
       FOR #Idx2 := 1 TO #Idx1 + 1 DO
           IF #ArrayTemp[#Idx2].Position > #MaxVal THEN
               #MaxVal := #ArrayTemp[#Idx2].Position;
               #MaxCarr := #ArrayTemp[#Idx2].CarrierNumber;
               #MaxIdx1 := #Idx2;
           END_IF;
       END_FOR;
       IF #MaxIdx1 > #Idx1 THEN
           #ArrayTemp[#MaxIdx1].Position := #ArrayTemp[#Idx1].Position;
           #ArrayTemp[#MaxIdx1].CarrierNumber := #ArrayTemp[#Idx1].CarrierNumber;
           #ArrayTemp[#Idx1].Position := #MaxVal;
           #ArrayTemp[#Idx1].CarrierNumber := #MaxCarr;

       END_IF;

   END_FOR;
   #ZonePositionArrayOut := #ArrayTemp;
END_FUNCTION

FUNCTION "FC107_FindLastZnPos" : Void   // FC107, SCL
{ S7_Optimized_Access := 'FALSE' }
VERSION : 0.1
   VAR_INPUT
      Zone : Int;
      TotalPosition : Int;
   END_VAR
   VAR_OUTPUT
      LastCarrierZnPos : Word;
   END_VAR
   VAR_TEMP
      ZnPosCounter : Int;
      ZoneFound : Word;
      CarrierCounter : Int;
      SortArrayIndex : Int;
      ArrayIndex : Int;
      Idx1 : Int;
      MaxVal : Int;
      MaxIdx1 : Int;
      Max : Int;
      Idx2 : Int;
      SelectionSort : Int;
   END_VAR
BEGIN
       #ZnPosCounter := #TotalPosition;
       WHILE #ZnPosCounter >= 1 DO

           IF "EMS".Zone[#Zone].CarrierZnStatus[#ZnPosCounter].CarrierNumber <> 0 THEN
               ;
               #LastCarrierZnPos := #ZnPosCounter;
               RETURN;
           END_IF;
           #ZnPosCounter := #ZnPosCounter - 1;
       END_WHILE;
END_FUNCTION

FUNCTION "FC108_FindCarrierZNPos" : Void   // FC108, SCL
{ S7_Optimized_Access := 'FALSE' }
VERSION : 0.1
   VAR_INPUT
      Carrier : Word;
      Zone : Int;
      TotalPosition : Int;
   END_VAR
   VAR_OUTPUT
      CarrierZnPos : Word;
   END_VAR
   VAR_TEMP
      ZnPosCounter : Int;
      ZoneFound : Word;
      CarrierCounter : Int;
      SortArrayIndex : Int;
      ArrayIndex : Int;
      Idx1 : Int;
      MaxVal : Int;
      MaxIdx1 : Int;
      Max : Int;
      Idx2 : Int;
      SelectionSort : Int;
   END_VAR
BEGIN
   //[***********************************************************************************NO EDITS*******************************************************************************************************]
   //FC204 - Find Carrier Zone Position
   //Single loop Counter finds which #Zone Position. Zone Position is determined BY Value OF Max Carriers defined in  #Carrier is located based on #Zone Start Position AND End Position AND
   //records the result in the system "EMS" DB FOR each Zone and the results stored in the EMS.Zone[Zone].CarrierZnStatus[1 thru Max Carriers in Zone].Carrier Number
   //***************************************************************************************************************************************************************************************************   

       #ZnPosCounter := 1;
       FOR #ZnPosCounter := 1 TO #TotalPosition DO
           ;
           IF "EMS".Zone[#Zone].CarrierZnStatus[#ZnPosCounter].CarrierNumber = #Carrier THEN;
               ;
               #CarrierZnPos := #ZnPosCounter;
           END_IF;
       END_FOR;
END_FUNCTION

FUNCTION "FC109_FindDuplicateCarrier" : Void   // FC109, SCL
{ S7_Optimized_Access := 'TRUE' }
VERSION : 0.1
   VAR_INPUT
      Carrier : Array[0..99] of "UDT_CarrierStructure";
      TotalCarriers : Int;
   END_VAR
   VAR_OUTPUT
      DuplicateFound : Bool;
      DuplicateCarrierNumber : Word;
      FirstDuplicatePosition : Word;
      SecondDuplicate : Word;
   END_VAR
   VAR_TEMP
      CarrierFindCnt : Int;
      temp1 : Int;
      CarrierCounter : Int;
      CarrierFindArray : Array[0..99] of "UDT_CarrierStructure";
   END_VAR
BEGIN
   //Sorts Carriers in Called Zone TO place in correct sequence within  Zone. Zones are divided into position based on MaxCarriers allowed in Zone as set in the Zone setup function block.


   #DuplicateFound := FALSE;
   #CarrierCounter := 1;
   #CarrierFindCnt := 1;
   #CarrierFindArray := #Carrier;
   FOR #CarrierFindCnt := 1 TO #TotalCarriers DO
       ;
       WHILE #CarrierCounter <= #TotalCarriers DO
           ;
           IF #Carrier[#CarrierCounter].SDC_IN.CarrierNumber = #CarrierFindArray[#CarrierFindCnt].SDC_IN.CarrierNumber AND #CarrierCounter <> #CarrierFindCnt AND #Carrier[#CarrierCounter].SDC_IN.CarrierNumber <> 0 THEN
               #DuplicateFound := TRUE;
               #FirstDuplicatePosition:= #Carrier[#CarrierCounter].SDC_IN.CarrierPosition;
               #SecondDuplicate := #Carrier[#CarrierFindCnt].SDC_IN.CarrierPosition;
               #DuplicateCarrierNumber := #CarrierFindArray[#CarrierFindCnt].SDC_IN.CarrierNumber;
               RETURN;
           END_IF;
           #CarrierCounter := #CarrierCounter + 1;
       END_WHILE;

       #CarrierCounter := 1;
   END_FOR;
END_FUNCTION

FUNCTION "FC110_HMIZonePosTracking" : Void   // FC110, SCL
{ S7_Optimized_Access := 'FALSE' }
VERSION : 0.1
   VAR_INPUT
      Zone : Int;
      TotalZones : Int;
      TotalCarriers : Int;
      MaxCarrierPosns : Int;
   END_VAR
   VAR_OUTPUT
      HMIZonePositionDisplay : Array[1..20] of "UDT_HMIZonePositionStructure";
   END_VAR
   VAR_TEMP
      PositionCounter : Int;
      ZoneFound : Word;
      CarrierCounter : Int;
      ZouneFound : Int;
   END_VAR
BEGIN

       FOR #PositionCounter := 1 TO #MaxCarrierPosns BY 1 DO
           FOR #CarrierCounter := 1 TO #TotalCarriers BY 1 DO
               ;
               IF "EMS".Carrier[#CarrierCounter].Position >= "EMS".Zone[#Zone].HMIZonePositions[#PositionCounter].ZonePosition AND
                   "EMS".Carrier[#CarrierCounter].Position < "EMS".Zone[#Zone].HMIZonePositions[#PositionCounter + 1].ZonePosition
               THEN
                   #HMIZonePositionDisplay[#PositionCounter].CarrierNumber := #CarrierCounter;
                   #HMIZonePositionDisplay[#PositionCounter].CarrierPosition := "EMS".Carrier[#CarrierCounter].Position;
                   #HMIZonePositionDisplay[#PositionCounter].Faulted := "EMS".Carrier[#CarrierCounter].Faulted;
                   EXIT;
               ELSE
                   ;
                   #HMIZonePositionDisplay[#PositionCounter].CarrierNumber := 0;
                   #HMIZonePositionDisplay[#PositionCounter].CarrierPosition := 0;
                   #HMIZonePositionDisplay[#PositionCounter].Faulted := 0;
               END_IF;
               "FC206CarrierLoop" := #CarrierCounter;
           END_FOR;
       "FC206PositionLoop" := #PositionCounter;
   END_FOR;
END_FUNCTION

FUNCTION "FC111_HMI_Status" : Void   // FC111, LAD
{ S7_Optimized_Access := 'TRUE' }
VERSION : 0.1
BEGIN

REGION Network 1
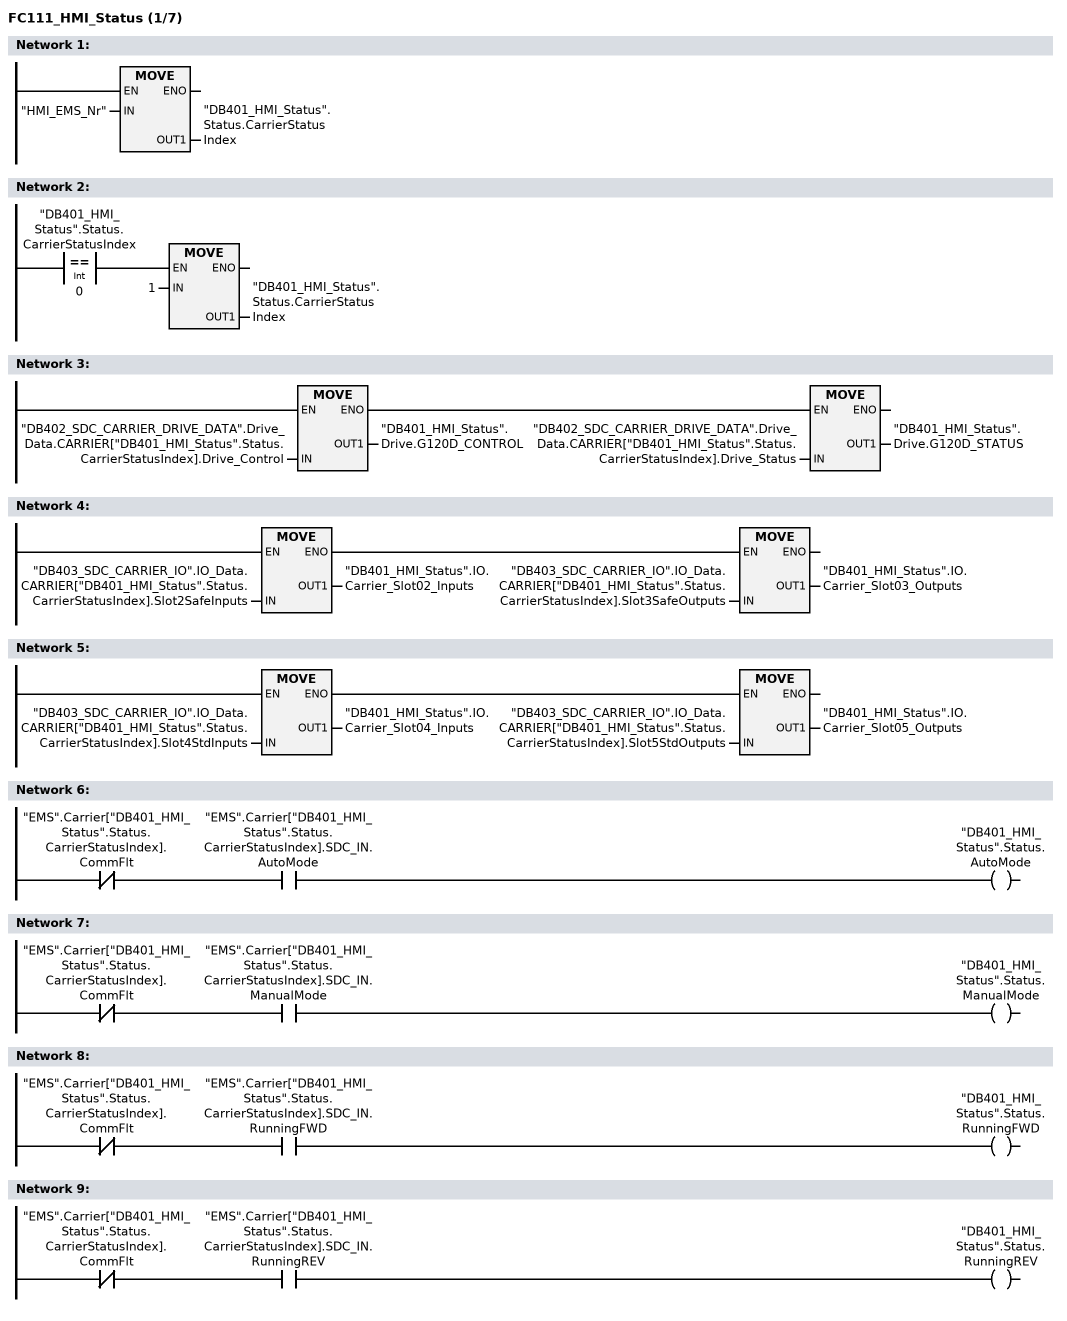
   RUNG wire#powerrail
      Move(in := "HMI_EMS_Nr", out1 => "DB401_HMI_Status".Status.CarrierStatusIndex)
   END_RUNG
   // the same network as SCL:
   "DB401_HMI_Status".Status.CarrierStatusIndex := "HMI_EMS_Nr";
END_REGION

REGION Network 2
   RUNG wire#powerrail
      { S7_Templates := "SrcType := Int" } EQ_Contact(in1 := "DB401_HMI_Status".Status.CarrierStatusIndex, in2 := 0)
      Move(in := 1, out1 => "DB401_HMI_Status".Status.CarrierStatusIndex)
   END_RUNG
   // the same network as SCL:
   IF "DB401_HMI_Status".Status.CarrierStatusIndex = 0 THEN
       "DB401_HMI_Status".Status.CarrierStatusIndex := 1;
   END_IF;
END_REGION

REGION Network 3
   RUNG wire#powerrail
      Move(in := "DB402_SDC_CARRIER_DRIVE_DATA".Drive_Data.CARRIER["DB401_HMI_Status".Status.CarrierStatusIndex].Drive_Control, out1 => "DB401_HMI_Status".Drive.G120D_CONTROL)
      Move(in := "DB402_SDC_CARRIER_DRIVE_DATA".Drive_Data.CARRIER["DB401_HMI_Status".Status.CarrierStatusIndex].Drive_Status, out1 => "DB401_HMI_Status".Drive.G120D_STATUS)
   END_RUNG
   // the same network as SCL:
   "DB401_HMI_Status".Drive.G120D_CONTROL := "DB402_SDC_CARRIER_DRIVE_DATA".Drive_Data.CARRIER["DB401_HMI_Status".Status.CarrierStatusIndex].Drive_Control;
   "DB401_HMI_Status".Drive.G120D_STATUS := "DB402_SDC_CARRIER_DRIVE_DATA".Drive_Data.CARRIER["DB401_HMI_Status".Status.CarrierStatusIndex].Drive_Status;
END_REGION

REGION Network 4
   RUNG wire#powerrail
      Move(in := "DB403_SDC_CARRIER_IO".IO_Data.CARRIER["DB401_HMI_Status".Status.CarrierStatusIndex].Slot2SafeInputs, out1 => "DB401_HMI_Status".IO.Carrier_Slot02_Inputs)
      Move(in := "DB403_SDC_CARRIER_IO".IO_Data.CARRIER["DB401_HMI_Status".Status.CarrierStatusIndex].Slot3SafeOutputs, out1 => "DB401_HMI_Status".IO.Carrier_Slot03_Outputs)
   END_RUNG
   // the same network as SCL:
   "DB401_HMI_Status".IO.Carrier_Slot02_Inputs := "DB403_SDC_CARRIER_IO".IO_Data.CARRIER["DB401_HMI_Status".Status.CarrierStatusIndex].Slot2SafeInputs;
   "DB401_HMI_Status".IO.Carrier_Slot03_Outputs := "DB403_SDC_CARRIER_IO".IO_Data.CARRIER["DB401_HMI_Status".Status.CarrierStatusIndex].Slot3SafeOutputs;
END_REGION

REGION Network 5
   RUNG wire#powerrail
      Move(in := "DB403_SDC_CARRIER_IO".IO_Data.CARRIER["DB401_HMI_Status".Status.CarrierStatusIndex].Slot4StdInputs, out1 => "DB401_HMI_Status".IO.Carrier_Slot04_Inputs)
      Move(in := "DB403_SDC_CARRIER_IO".IO_Data.CARRIER["DB401_HMI_Status".Status.CarrierStatusIndex].Slot5StdOutputs, out1 => "DB401_HMI_Status".IO.Carrier_Slot05_Outputs)
   END_RUNG
   // the same network as SCL:
   "DB401_HMI_Status".IO.Carrier_Slot04_Inputs := "DB403_SDC_CARRIER_IO".IO_Data.CARRIER["DB401_HMI_Status".Status.CarrierStatusIndex].Slot4StdInputs;
   "DB401_HMI_Status".IO.Carrier_Slot05_Outputs := "DB403_SDC_CARRIER_IO".IO_Data.CARRIER["DB401_HMI_Status".Status.CarrierStatusIndex].Slot5StdOutputs;
END_REGION

REGION Network 6
   RUNG wire#powerrail
      I_Contact( "EMS".Carrier["DB401_HMI_Status".Status.CarrierStatusIndex].CommFlt )
      Contact( "EMS".Carrier["DB401_HMI_Status".Status.CarrierStatusIndex].SDC_IN.AutoMode )
      Coil( "DB401_HMI_Status".Status.AutoMode )
   END_RUNG
   // the same network as SCL:
   "DB401_HMI_Status".Status.AutoMode := NOT "EMS".Carrier["DB401_HMI_Status".Status.CarrierStatusIndex].CommFlt AND "EMS".Carrier["DB401_HMI_Status".Status.CarrierStatusIndex].SDC_IN.AutoMode;
END_REGION

REGION Network 7
   RUNG wire#powerrail
      I_Contact( "EMS".Carrier["DB401_HMI_Status".Status.CarrierStatusIndex].CommFlt )
      Contact( "EMS".Carrier["DB401_HMI_Status".Status.CarrierStatusIndex].SDC_IN.ManualMode )
      Coil( "DB401_HMI_Status".Status.ManualMode )
   END_RUNG
   // the same network as SCL:
   "DB401_HMI_Status".Status.ManualMode := NOT "EMS".Carrier["DB401_HMI_Status".Status.CarrierStatusIndex].CommFlt AND "EMS".Carrier["DB401_HMI_Status".Status.CarrierStatusIndex].SDC_IN.ManualMode;
END_REGION

REGION Network 8
   RUNG wire#powerrail
      I_Contact( "EMS".Carrier["DB401_HMI_Status".Status.CarrierStatusIndex].CommFlt )
      Contact( "EMS".Carrier["DB401_HMI_Status".Status.CarrierStatusIndex].SDC_IN.RunningFWD )
      Coil( "DB401_HMI_Status".Status.RunningFWD )
   END_RUNG
   // the same network as SCL:
   "DB401_HMI_Status".Status.RunningFWD := NOT "EMS".Carrier["DB401_HMI_Status".Status.CarrierStatusIndex].CommFlt AND "EMS".Carrier["DB401_HMI_Status".Status.CarrierStatusIndex].SDC_IN.RunningFWD;
END_REGION

REGION Network 9
   RUNG wire#powerrail
      I_Contact( "EMS".Carrier["DB401_HMI_Status".Status.CarrierStatusIndex].CommFlt )
      Contact( "EMS".Carrier["DB401_HMI_Status".Status.CarrierStatusIndex].SDC_IN.RunningREV )
      Coil( "DB401_HMI_Status".Status.RunningREV )
   END_RUNG
   // the same network as SCL:
   "DB401_HMI_Status".Status.RunningREV := NOT "EMS".Carrier["DB401_HMI_Status".Status.CarrierStatusIndex].CommFlt AND "EMS".Carrier["DB401_HMI_Status".Status.CarrierStatusIndex].SDC_IN.RunningREV;
END_REGION

REGION Network 10
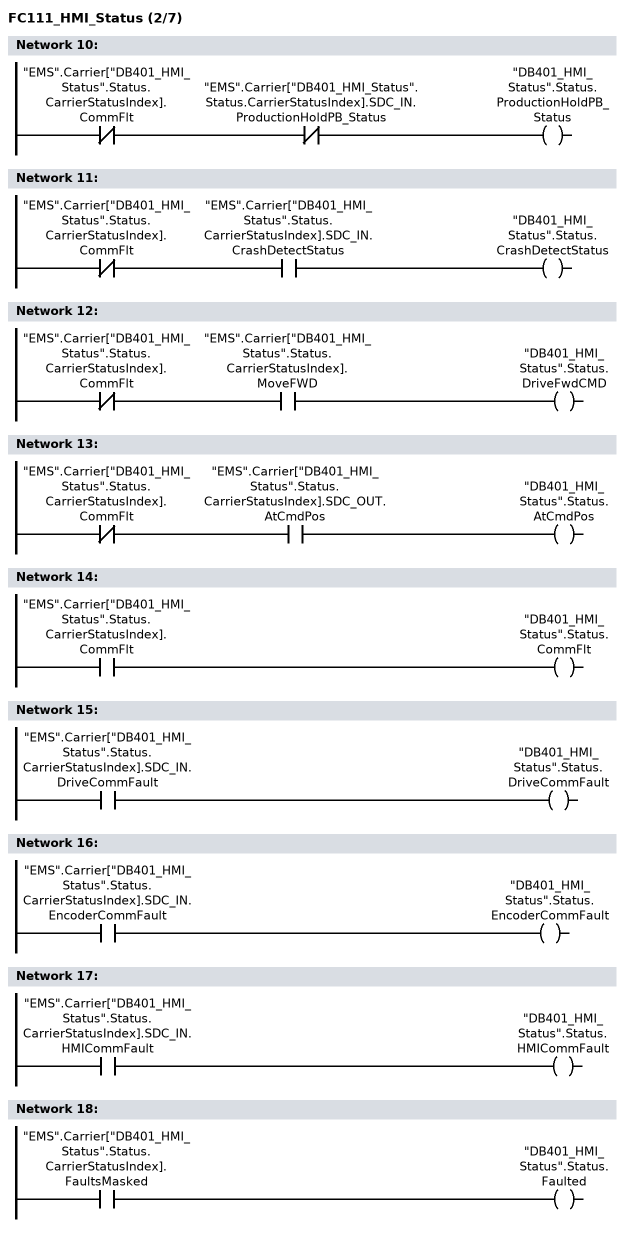
   RUNG wire#powerrail
      I_Contact( "EMS".Carrier["DB401_HMI_Status".Status.CarrierStatusIndex].CommFlt )
      I_Contact( "EMS".Carrier["DB401_HMI_Status".Status.CarrierStatusIndex].SDC_IN.ProductionHoldPB_Status )
      Coil( "DB401_HMI_Status".Status.ProductionHoldPB_Status )
   END_RUNG
   // the same network as SCL:
   "DB401_HMI_Status".Status.ProductionHoldPB_Status := NOT "EMS".Carrier["DB401_HMI_Status".Status.CarrierStatusIndex].CommFlt AND NOT "EMS".Carrier["DB401_HMI_Status".Status.CarrierStatusIndex].SDC_IN.ProductionHoldPB_Status;
END_REGION

REGION Network 11
   RUNG wire#powerrail
      I_Contact( "EMS".Carrier["DB401_HMI_Status".Status.CarrierStatusIndex].CommFlt )
      Contact( "EMS".Carrier["DB401_HMI_Status".Status.CarrierStatusIndex].SDC_IN.CrashDetectStatus )
      Coil( "DB401_HMI_Status".Status.CrashDetectStatus )
   END_RUNG
   // the same network as SCL:
   "DB401_HMI_Status".Status.CrashDetectStatus := NOT "EMS".Carrier["DB401_HMI_Status".Status.CarrierStatusIndex].CommFlt AND "EMS".Carrier["DB401_HMI_Status".Status.CarrierStatusIndex].SDC_IN.CrashDetectStatus;
END_REGION

REGION Network 12
   RUNG wire#powerrail
      I_Contact( "EMS".Carrier["DB401_HMI_Status".Status.CarrierStatusIndex].CommFlt )
      Contact( "EMS".Carrier["DB401_HMI_Status".Status.CarrierStatusIndex].MoveFWD )
      Coil( "DB401_HMI_Status".Status.DriveFwdCMD )
   END_RUNG
   // the same network as SCL:
   "DB401_HMI_Status".Status.DriveFwdCMD := NOT "EMS".Carrier["DB401_HMI_Status".Status.CarrierStatusIndex].CommFlt AND "EMS".Carrier["DB401_HMI_Status".Status.CarrierStatusIndex].MoveFWD;
END_REGION

REGION Network 13
   RUNG wire#powerrail
      I_Contact( "EMS".Carrier["DB401_HMI_Status".Status.CarrierStatusIndex].CommFlt )
      Contact( "EMS".Carrier["DB401_HMI_Status".Status.CarrierStatusIndex].SDC_OUT.AtCmdPos )
      Coil( "DB401_HMI_Status".Status.AtCmdPos )
   END_RUNG
   // the same network as SCL:
   "DB401_HMI_Status".Status.AtCmdPos := NOT "EMS".Carrier["DB401_HMI_Status".Status.CarrierStatusIndex].CommFlt AND "EMS".Carrier["DB401_HMI_Status".Status.CarrierStatusIndex].SDC_OUT.AtCmdPos;
END_REGION

REGION Network 14
   RUNG wire#powerrail
      Contact( "EMS".Carrier["DB401_HMI_Status".Status.CarrierStatusIndex].CommFlt )
      Coil( "DB401_HMI_Status".Status.CommFlt )
   END_RUNG
   // the same network as SCL:
   "DB401_HMI_Status".Status.CommFlt := "EMS".Carrier["DB401_HMI_Status".Status.CarrierStatusIndex].CommFlt;
END_REGION

REGION Network 15
   RUNG wire#powerrail
      Contact( "EMS".Carrier["DB401_HMI_Status".Status.CarrierStatusIndex].SDC_IN.DriveCommFault )
      Coil( "DB401_HMI_Status".Status.DriveCommFault )
   END_RUNG
   // the same network as SCL:
   "DB401_HMI_Status".Status.DriveCommFault := "EMS".Carrier["DB401_HMI_Status".Status.CarrierStatusIndex].SDC_IN.DriveCommFault;
END_REGION

REGION Network 16
   RUNG wire#powerrail
      Contact( "EMS".Carrier["DB401_HMI_Status".Status.CarrierStatusIndex].SDC_IN.EncoderCommFault )
      Coil( "DB401_HMI_Status".Status.EncoderCommFault )
   END_RUNG
   // the same network as SCL:
   "DB401_HMI_Status".Status.EncoderCommFault := "EMS".Carrier["DB401_HMI_Status".Status.CarrierStatusIndex].SDC_IN.EncoderCommFault;
END_REGION

REGION Network 17
   RUNG wire#powerrail
      Contact( "EMS".Carrier["DB401_HMI_Status".Status.CarrierStatusIndex].SDC_IN.HMICommFault )
      Coil( "DB401_HMI_Status".Status.HMICommFault )
   END_RUNG
   // the same network as SCL:
   "DB401_HMI_Status".Status.HMICommFault := "EMS".Carrier["DB401_HMI_Status".Status.CarrierStatusIndex].SDC_IN.HMICommFault;
END_REGION

REGION Network 18
   RUNG wire#powerrail
      Contact( "EMS".Carrier["DB401_HMI_Status".Status.CarrierStatusIndex].FaultsMasked )
      Coil( "DB401_HMI_Status".Status.Faulted )
   END_RUNG
   // the same network as SCL:
   "DB401_HMI_Status".Status.Faulted := "EMS".Carrier["DB401_HMI_Status".Status.CarrierStatusIndex].FaultsMasked;
END_REGION

REGION Network 19: PRODUCTION STOP WARNING 'H07'
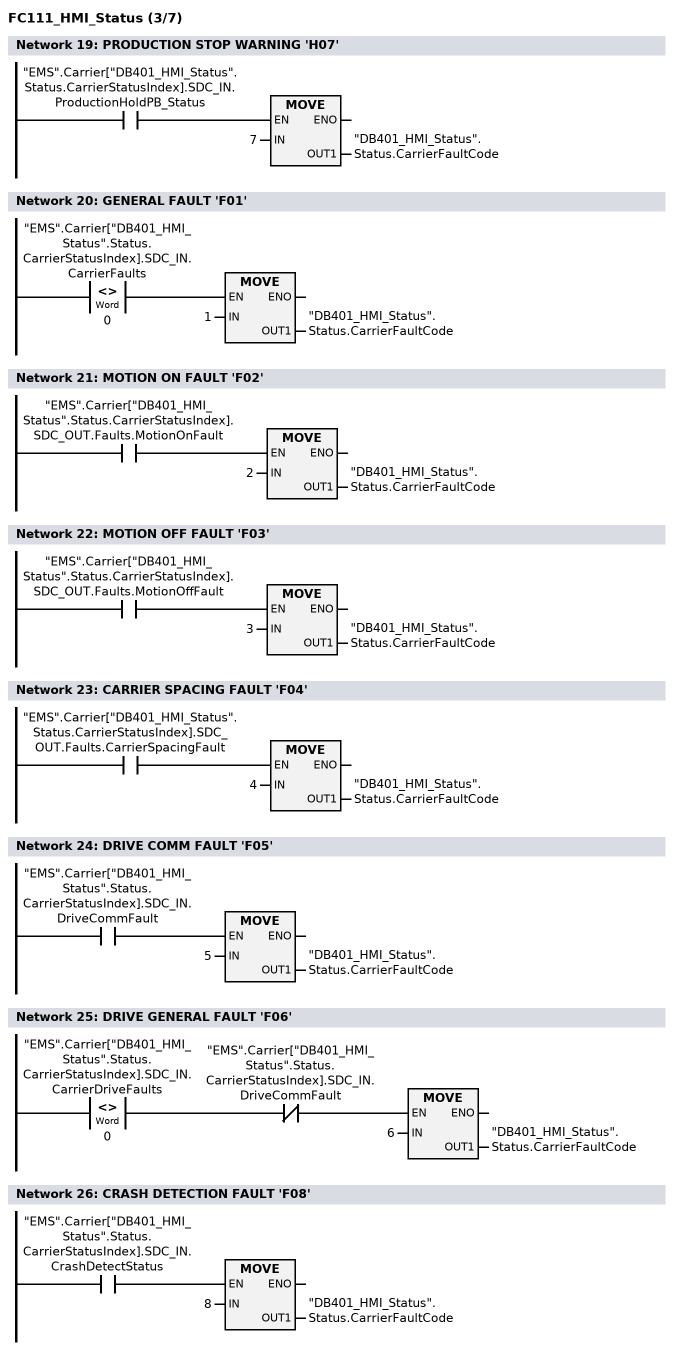
   RUNG wire#powerrail
      Contact( "EMS".Carrier["DB401_HMI_Status".Status.CarrierStatusIndex].SDC_IN.ProductionHoldPB_Status )
      Move(in := 7, out1 => "DB401_HMI_Status".Status.CarrierFaultCode)
   END_RUNG
   // the same network as SCL:
   IF "EMS".Carrier["DB401_HMI_Status".Status.CarrierStatusIndex].SDC_IN.ProductionHoldPB_Status THEN
       "DB401_HMI_Status".Status.CarrierFaultCode := 7;
   END_IF;
END_REGION

REGION Network 20: GENERAL FAULT 'F01'
   RUNG wire#powerrail
      { S7_Templates := "SrcType := Word" } NE_Contact(in1 := "EMS".Carrier["DB401_HMI_Status".Status.CarrierStatusIndex].SDC_IN.CarrierFaults, in2 := 0)
      Move(in := 1, out1 => "DB401_HMI_Status".Status.CarrierFaultCode)
   END_RUNG
   // the same network as SCL:
   IF "EMS".Carrier["DB401_HMI_Status".Status.CarrierStatusIndex].SDC_IN.CarrierFaults <> 0 THEN
       "DB401_HMI_Status".Status.CarrierFaultCode := 1;
   END_IF;
END_REGION

REGION Network 21: MOTION ON FAULT 'F02'
   RUNG wire#powerrail
      Contact( "EMS".Carrier["DB401_HMI_Status".Status.CarrierStatusIndex].SDC_OUT.Faults.MotionOnFault )
      Move(in := 2, out1 => "DB401_HMI_Status".Status.CarrierFaultCode)
   END_RUNG
   // the same network as SCL:
   IF "EMS".Carrier["DB401_HMI_Status".Status.CarrierStatusIndex].SDC_OUT.Faults.MotionOnFault THEN
       "DB401_HMI_Status".Status.CarrierFaultCode := 2;
   END_IF;
END_REGION

REGION Network 22: MOTION OFF FAULT 'F03'
   RUNG wire#powerrail
      Contact( "EMS".Carrier["DB401_HMI_Status".Status.CarrierStatusIndex].SDC_OUT.Faults.MotionOffFault )
      Move(in := 3, out1 => "DB401_HMI_Status".Status.CarrierFaultCode)
   END_RUNG
   // the same network as SCL:
   IF "EMS".Carrier["DB401_HMI_Status".Status.CarrierStatusIndex].SDC_OUT.Faults.MotionOffFault THEN
       "DB401_HMI_Status".Status.CarrierFaultCode := 3;
   END_IF;
END_REGION

REGION Network 23: CARRIER SPACING FAULT 'F04'
   RUNG wire#powerrail
      Contact( "EMS".Carrier["DB401_HMI_Status".Status.CarrierStatusIndex].SDC_OUT.Faults.CarrierSpacingFault )
      Move(in := 4, out1 => "DB401_HMI_Status".Status.CarrierFaultCode)
   END_RUNG
   // the same network as SCL:
   IF "EMS".Carrier["DB401_HMI_Status".Status.CarrierStatusIndex].SDC_OUT.Faults.CarrierSpacingFault THEN
       "DB401_HMI_Status".Status.CarrierFaultCode := 4;
   END_IF;
END_REGION

REGION Network 24: DRIVE COMM FAULT 'F05'
   RUNG wire#powerrail
      Contact( "EMS".Carrier["DB401_HMI_Status".Status.CarrierStatusIndex].SDC_IN.DriveCommFault )
      Move(in := 5, out1 => "DB401_HMI_Status".Status.CarrierFaultCode)
   END_RUNG
   // the same network as SCL:
   IF "EMS".Carrier["DB401_HMI_Status".Status.CarrierStatusIndex].SDC_IN.DriveCommFault THEN
       "DB401_HMI_Status".Status.CarrierFaultCode := 5;
   END_IF;
END_REGION

REGION Network 25: DRIVE GENERAL FAULT 'F06'
   RUNG wire#powerrail
      { S7_Templates := "SrcType := Word" } NE_Contact(in1 := "EMS".Carrier["DB401_HMI_Status".Status.CarrierStatusIndex].SDC_IN.CarrierDriveFaults, in2 := 0)
      I_Contact( "EMS".Carrier["DB401_HMI_Status".Status.CarrierStatusIndex].SDC_IN.DriveCommFault )
      Move(in := 6, out1 => "DB401_HMI_Status".Status.CarrierFaultCode)
   END_RUNG
   // the same network as SCL:
   IF ("EMS".Carrier["DB401_HMI_Status".Status.CarrierStatusIndex].SDC_IN.CarrierDriveFaults <> 0) AND NOT "EMS".Carrier["DB401_HMI_Status".Status.CarrierStatusIndex].SDC_IN.DriveCommFault THEN
       "DB401_HMI_Status".Status.CarrierFaultCode := 6;
   END_IF;
END_REGION

REGION Network 26: CRASH DETECTION FAULT 'F08'
   RUNG wire#powerrail
      Contact( "EMS".Carrier["DB401_HMI_Status".Status.CarrierStatusIndex].SDC_IN.CrashDetectStatus )
      Move(in := 8, out1 => "DB401_HMI_Status".Status.CarrierFaultCode)
   END_RUNG
   // the same network as SCL:
   IF "EMS".Carrier["DB401_HMI_Status".Status.CarrierStatusIndex].SDC_IN.CrashDetectStatus THEN
       "DB401_HMI_Status".Status.CarrierFaultCode := 8;
   END_IF;
END_REGION

REGION Network 27: DRIVE ERROR INTERNAL COMM FAULT 'F15'
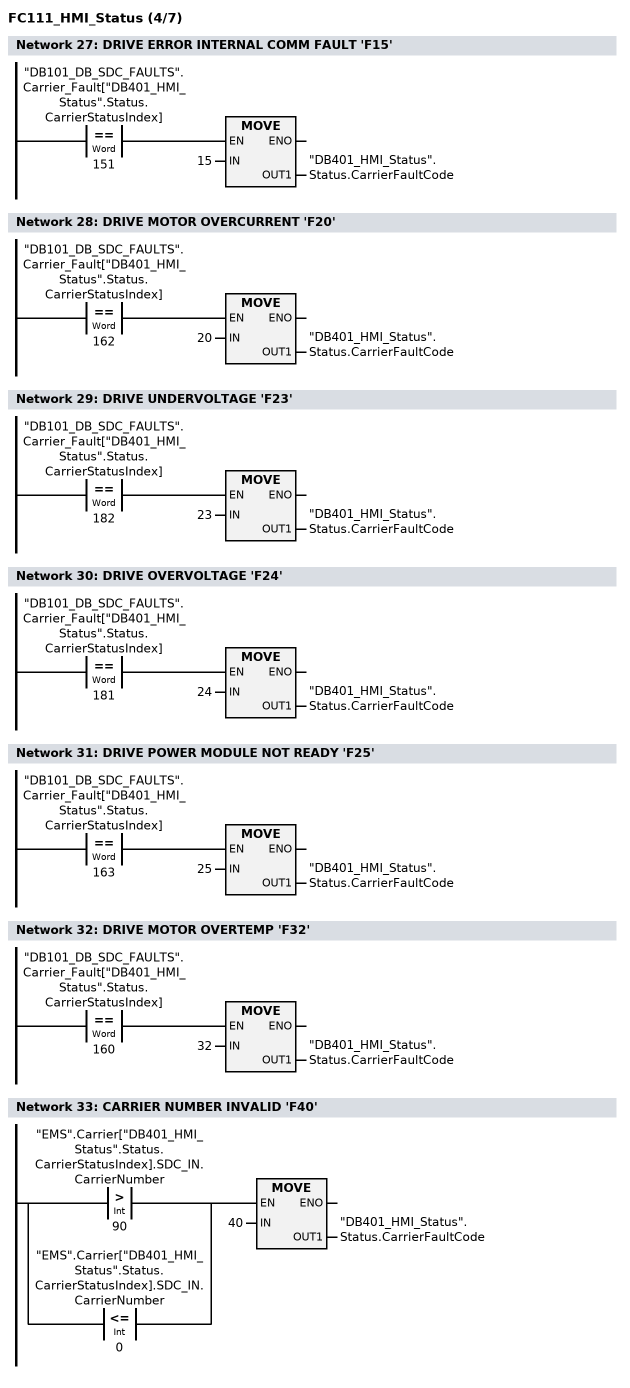
   RUNG wire#powerrail
      { S7_Templates := "SrcType := Word" } EQ_Contact(in1 := "DB101_DB_SDC_FAULTS".Carrier_Fault["DB401_HMI_Status".Status.CarrierStatusIndex], in2 := 151)
      Move(in := 15, out1 => "DB401_HMI_Status".Status.CarrierFaultCode)
   END_RUNG
   // the same network as SCL:
   IF "DB101_DB_SDC_FAULTS".Carrier_Fault["DB401_HMI_Status".Status.CarrierStatusIndex] = 151 THEN
       "DB401_HMI_Status".Status.CarrierFaultCode := 15;
   END_IF;
END_REGION

REGION Network 28: DRIVE MOTOR OVERCURRENT 'F20'
   RUNG wire#powerrail
      { S7_Templates := "SrcType := Word" } EQ_Contact(in1 := "DB101_DB_SDC_FAULTS".Carrier_Fault["DB401_HMI_Status".Status.CarrierStatusIndex], in2 := 162)
      Move(in := 20, out1 => "DB401_HMI_Status".Status.CarrierFaultCode)
   END_RUNG
   // the same network as SCL:
   IF "DB101_DB_SDC_FAULTS".Carrier_Fault["DB401_HMI_Status".Status.CarrierStatusIndex] = 162 THEN
       "DB401_HMI_Status".Status.CarrierFaultCode := 20;
   END_IF;
END_REGION

REGION Network 29: DRIVE UNDERVOLTAGE 'F23'
   RUNG wire#powerrail
      { S7_Templates := "SrcType := Word" } EQ_Contact(in1 := "DB101_DB_SDC_FAULTS".Carrier_Fault["DB401_HMI_Status".Status.CarrierStatusIndex], in2 := 182)
      Move(in := 23, out1 => "DB401_HMI_Status".Status.CarrierFaultCode)
   END_RUNG
   // the same network as SCL:
   IF "DB101_DB_SDC_FAULTS".Carrier_Fault["DB401_HMI_Status".Status.CarrierStatusIndex] = 182 THEN
       "DB401_HMI_Status".Status.CarrierFaultCode := 23;
   END_IF;
END_REGION

REGION Network 30: DRIVE OVERVOLTAGE 'F24'
   RUNG wire#powerrail
      { S7_Templates := "SrcType := Word" } EQ_Contact(in1 := "DB101_DB_SDC_FAULTS".Carrier_Fault["DB401_HMI_Status".Status.CarrierStatusIndex], in2 := 181)
      Move(in := 24, out1 => "DB401_HMI_Status".Status.CarrierFaultCode)
   END_RUNG
   // the same network as SCL:
   IF "DB101_DB_SDC_FAULTS".Carrier_Fault["DB401_HMI_Status".Status.CarrierStatusIndex] = 181 THEN
       "DB401_HMI_Status".Status.CarrierFaultCode := 24;
   END_IF;
END_REGION

REGION Network 31: DRIVE POWER MODULE NOT READY 'F25'
   RUNG wire#powerrail
      { S7_Templates := "SrcType := Word" } EQ_Contact(in1 := "DB101_DB_SDC_FAULTS".Carrier_Fault["DB401_HMI_Status".Status.CarrierStatusIndex], in2 := 163)
      Move(in := 25, out1 => "DB401_HMI_Status".Status.CarrierFaultCode)
   END_RUNG
   // the same network as SCL:
   IF "DB101_DB_SDC_FAULTS".Carrier_Fault["DB401_HMI_Status".Status.CarrierStatusIndex] = 163 THEN
       "DB401_HMI_Status".Status.CarrierFaultCode := 25;
   END_IF;
END_REGION

REGION Network 32: DRIVE MOTOR OVERTEMP 'F32'
   RUNG wire#powerrail
      { S7_Templates := "SrcType := Word" } EQ_Contact(in1 := "DB101_DB_SDC_FAULTS".Carrier_Fault["DB401_HMI_Status".Status.CarrierStatusIndex], in2 := 160)
      Move(in := 32, out1 => "DB401_HMI_Status".Status.CarrierFaultCode)
   END_RUNG
   // the same network as SCL:
   IF "DB101_DB_SDC_FAULTS".Carrier_Fault["DB401_HMI_Status".Status.CarrierStatusIndex] = 160 THEN
       "DB401_HMI_Status".Status.CarrierFaultCode := 32;
   END_IF;
END_REGION

REGION Network 33: CARRIER NUMBER INVALID 'F40'
   RUNG wire#powerrail
      { S7_Templates := "SrcType := Int" } GT_Contact(in1 := "EMS".Carrier["DB401_HMI_Status".Status.CarrierStatusIndex].SDC_IN.CarrierNumber, in2 := 90)
      wire#w1
      Move(in := 40, out1 => "DB401_HMI_Status".Status.CarrierFaultCode)
   END_RUNG
   RUNG wire#powerrail
      { S7_Templates := "SrcType := Int" } LE_Contact(in1 := "EMS".Carrier["DB401_HMI_Status".Status.CarrierStatusIndex].SDC_IN.CarrierNumber, in2 := 0)
   END_RUNG wire#w1
   // the same network as SCL:
   IF ("EMS".Carrier["DB401_HMI_Status".Status.CarrierStatusIndex].SDC_IN.CarrierNumber > 90) OR ("EMS".Carrier["DB401_HMI_Status".Status.CarrierStatusIndex].SDC_IN.CarrierNumber <= 0) THEN
       "DB401_HMI_Status".Status.CarrierFaultCode := 40;
   END_IF;
END_REGION

REGION Network 34: ENCODER FAULT 'F60'
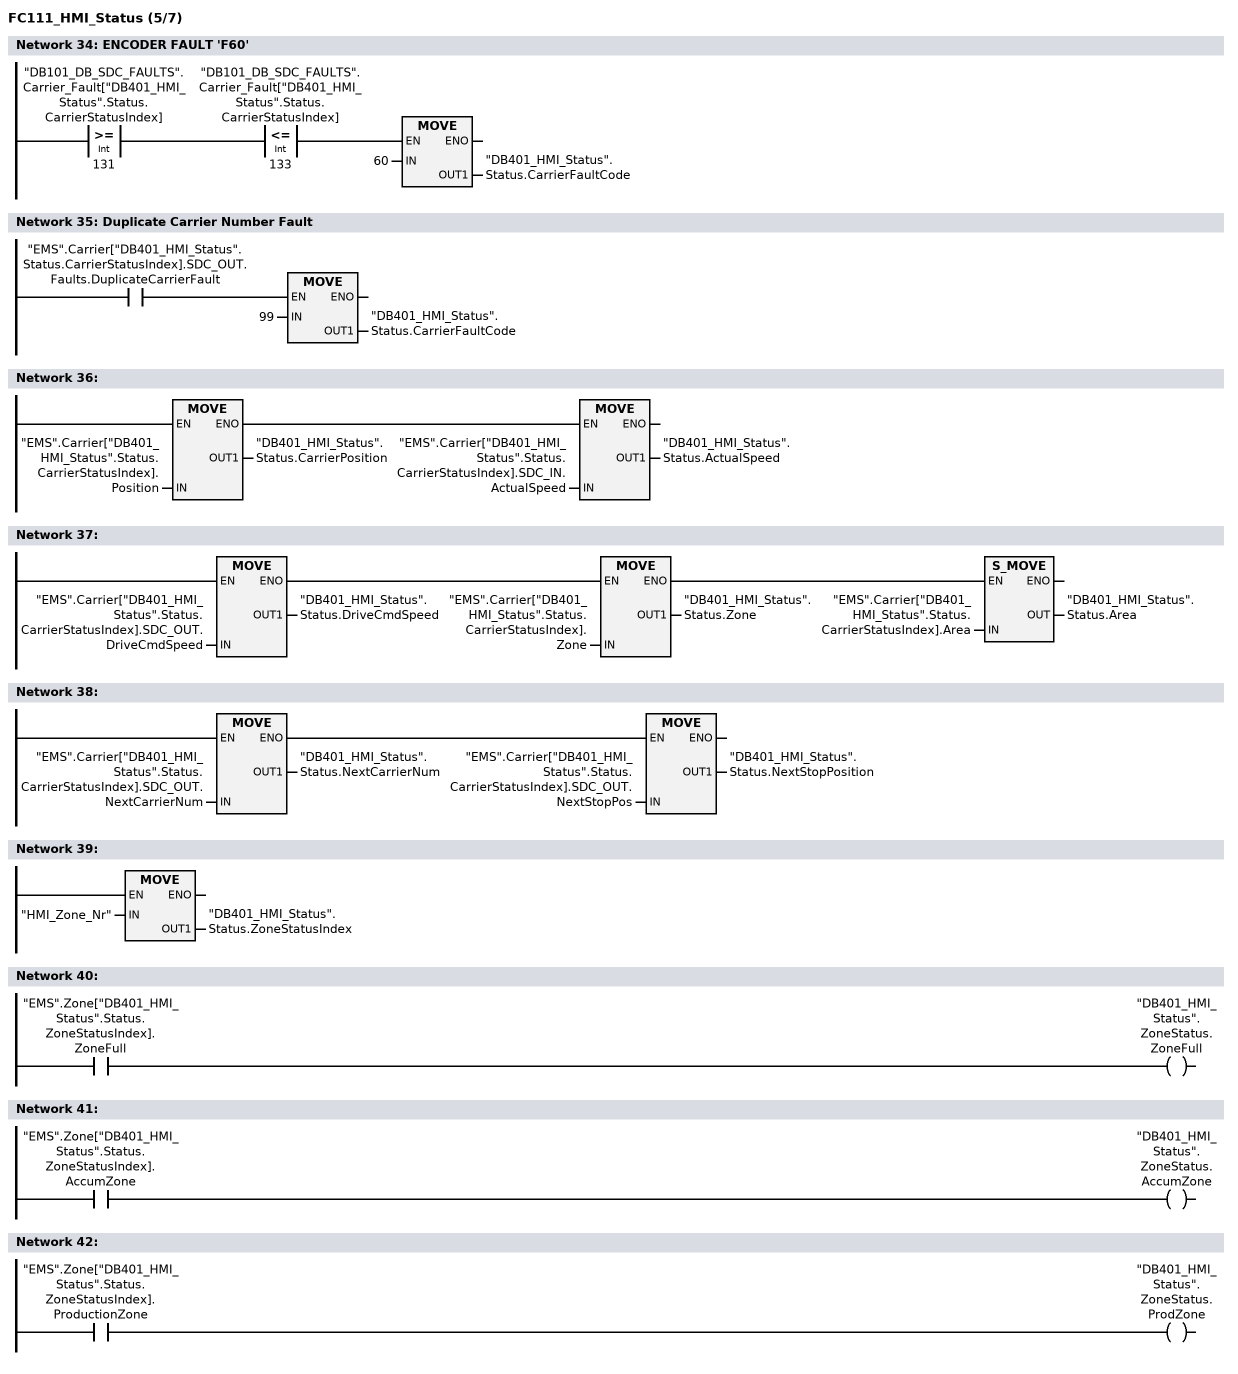
   RUNG wire#powerrail
      { S7_Templates := "SrcType := Int" } GE_Contact(in1 := "DB101_DB_SDC_FAULTS".Carrier_Fault["DB401_HMI_Status".Status.CarrierStatusIndex], in2 := 131)
      { S7_Templates := "SrcType := Int" } LE_Contact(in1 := "DB101_DB_SDC_FAULTS".Carrier_Fault["DB401_HMI_Status".Status.CarrierStatusIndex], in2 := 133)
      Move(in := 60, out1 => "DB401_HMI_Status".Status.CarrierFaultCode)
   END_RUNG
   // the same network as SCL:
   IF ("DB101_DB_SDC_FAULTS".Carrier_Fault["DB401_HMI_Status".Status.CarrierStatusIndex] >= 131) AND ("DB101_DB_SDC_FAULTS".Carrier_Fault["DB401_HMI_Status".Status.CarrierStatusIndex] <= 133) THEN
       "DB401_HMI_Status".Status.CarrierFaultCode := 60;
   END_IF;
END_REGION

REGION Network 35: Duplicate Carrier Number Fault
   RUNG wire#powerrail
      Contact( "EMS".Carrier["DB401_HMI_Status".Status.CarrierStatusIndex].SDC_OUT.Faults.DuplicateCarrierFault )
      Move(in := 99, out1 => "DB401_HMI_Status".Status.CarrierFaultCode)
   END_RUNG
   // the same network as SCL:
   IF "EMS".Carrier["DB401_HMI_Status".Status.CarrierStatusIndex].SDC_OUT.Faults.DuplicateCarrierFault THEN
       "DB401_HMI_Status".Status.CarrierFaultCode := 99;
   END_IF;
END_REGION

REGION Network 36
   RUNG wire#powerrail
      Move(in := "EMS".Carrier["DB401_HMI_Status".Status.CarrierStatusIndex].Position, out1 => "DB401_HMI_Status".Status.CarrierPosition)
      Move(in := "EMS".Carrier["DB401_HMI_Status".Status.CarrierStatusIndex].SDC_IN.ActualSpeed, out1 => "DB401_HMI_Status".Status.ActualSpeed)
   END_RUNG
   // the same network as SCL:
   "DB401_HMI_Status".Status.CarrierPosition := "EMS".Carrier["DB401_HMI_Status".Status.CarrierStatusIndex].Position;
   "DB401_HMI_Status".Status.ActualSpeed := "EMS".Carrier["DB401_HMI_Status".Status.CarrierStatusIndex].SDC_IN.ActualSpeed;
END_REGION

REGION Network 37
   RUNG wire#powerrail
      Move(in := "EMS".Carrier["DB401_HMI_Status".Status.CarrierStatusIndex].SDC_OUT.DriveCmdSpeed, out1 => "DB401_HMI_Status".Status.DriveCmdSpeed)
      Move(in := "EMS".Carrier["DB401_HMI_Status".Status.CarrierStatusIndex].Zone, out1 => "DB401_HMI_Status".Status.Zone)
      S_Move(in := "EMS".Carrier["DB401_HMI_Status".Status.CarrierStatusIndex].Area, out => "DB401_HMI_Status".Status.Area)
   END_RUNG
   // the same network as SCL:
   "DB401_HMI_Status".Status.DriveCmdSpeed := "EMS".Carrier["DB401_HMI_Status".Status.CarrierStatusIndex].SDC_OUT.DriveCmdSpeed;
   "DB401_HMI_Status".Status.Zone := "EMS".Carrier["DB401_HMI_Status".Status.CarrierStatusIndex].Zone;
   "DB401_HMI_Status".Status.Area := "EMS".Carrier["DB401_HMI_Status".Status.CarrierStatusIndex].Area;
END_REGION

REGION Network 38
   RUNG wire#powerrail
      Move(in := "EMS".Carrier["DB401_HMI_Status".Status.CarrierStatusIndex].SDC_OUT.NextCarrierNum, out1 => "DB401_HMI_Status".Status.NextCarrierNum)
      Move(in := "EMS".Carrier["DB401_HMI_Status".Status.CarrierStatusIndex].SDC_OUT.NextStopPos, out1 => "DB401_HMI_Status".Status.NextStopPosition)
   END_RUNG
   // the same network as SCL:
   "DB401_HMI_Status".Status.NextCarrierNum := "EMS".Carrier["DB401_HMI_Status".Status.CarrierStatusIndex].SDC_OUT.NextCarrierNum;
   "DB401_HMI_Status".Status.NextStopPosition := "EMS".Carrier["DB401_HMI_Status".Status.CarrierStatusIndex].SDC_OUT.NextStopPos;
END_REGION

REGION Network 39
   RUNG wire#powerrail
      Move(in := "HMI_Zone_Nr", out1 => "DB401_HMI_Status".Status.ZoneStatusIndex)
   END_RUNG
   // the same network as SCL:
   "DB401_HMI_Status".Status.ZoneStatusIndex := "HMI_Zone_Nr";
END_REGION

REGION Network 40
   RUNG wire#powerrail
      Contact( "EMS".Zone["DB401_HMI_Status".Status.ZoneStatusIndex].ZoneFull )
      Coil( "DB401_HMI_Status".ZoneStatus.ZoneFull )
   END_RUNG
   // the same network as SCL:
   "DB401_HMI_Status".ZoneStatus.ZoneFull := "EMS".Zone["DB401_HMI_Status".Status.ZoneStatusIndex].ZoneFull;
END_REGION

REGION Network 41
   RUNG wire#powerrail
      Contact( "EMS".Zone["DB401_HMI_Status".Status.ZoneStatusIndex].AccumZone )
      Coil( "DB401_HMI_Status".ZoneStatus.AccumZone )
   END_RUNG
   // the same network as SCL:
   "DB401_HMI_Status".ZoneStatus.AccumZone := "EMS".Zone["DB401_HMI_Status".Status.ZoneStatusIndex].AccumZone;
END_REGION

REGION Network 42
   RUNG wire#powerrail
      Contact( "EMS".Zone["DB401_HMI_Status".Status.ZoneStatusIndex].ProductionZone )
      Coil( "DB401_HMI_Status".ZoneStatus.ProdZone )
   END_RUNG
   // the same network as SCL:
   "DB401_HMI_Status".ZoneStatus.ProdZone := "EMS".Zone["DB401_HMI_Status".Status.ZoneStatusIndex].ProductionZone;
END_REGION

REGION Network 43
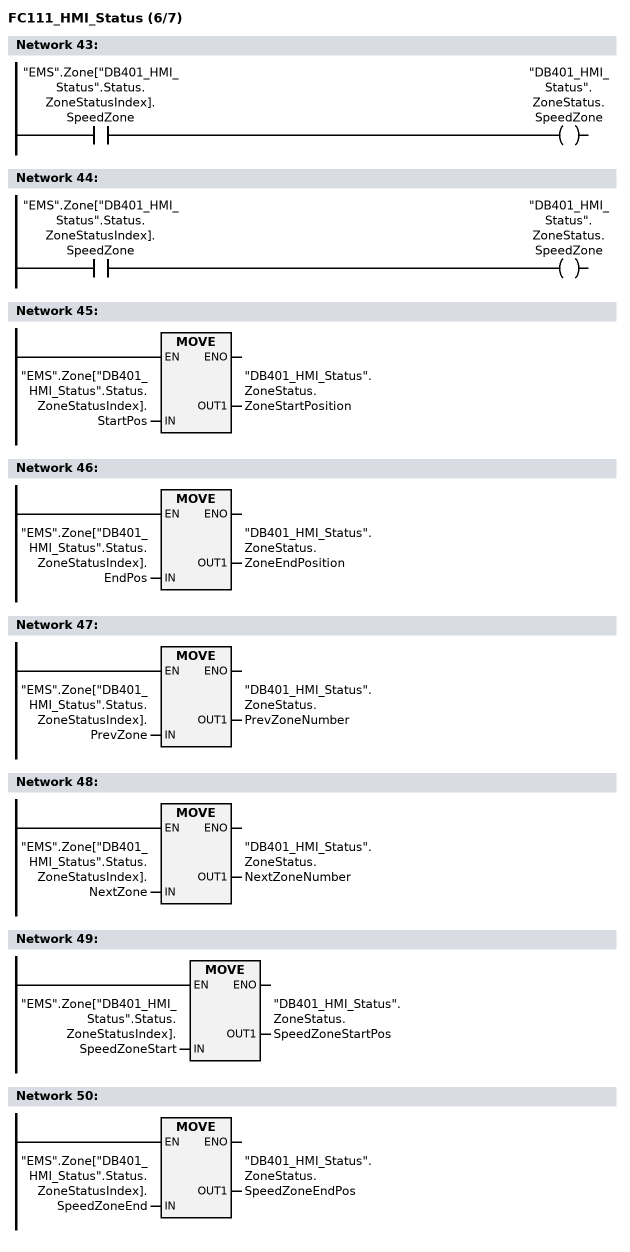
   RUNG wire#powerrail
      Contact( "EMS".Zone["DB401_HMI_Status".Status.ZoneStatusIndex].SpeedZone )
      Coil( "DB401_HMI_Status".ZoneStatus.SpeedZone )
   END_RUNG
   // the same network as SCL:
   "DB401_HMI_Status".ZoneStatus.SpeedZone := "EMS".Zone["DB401_HMI_Status".Status.ZoneStatusIndex].SpeedZone;
END_REGION

REGION Network 44
   RUNG wire#powerrail
      Contact( "EMS".Zone["DB401_HMI_Status".Status.ZoneStatusIndex].SpeedZone )
      Coil( "DB401_HMI_Status".ZoneStatus.SpeedZone )
   END_RUNG
   // the same network as SCL:
   "DB401_HMI_Status".ZoneStatus.SpeedZone := "EMS".Zone["DB401_HMI_Status".Status.ZoneStatusIndex].SpeedZone;
END_REGION

REGION Network 45
   RUNG wire#powerrail
      Move(in := "EMS".Zone["DB401_HMI_Status".Status.ZoneStatusIndex].StartPos, out1 => "DB401_HMI_Status".ZoneStatus.ZoneStartPosition)
   END_RUNG
   // the same network as SCL:
   "DB401_HMI_Status".ZoneStatus.ZoneStartPosition := "EMS".Zone["DB401_HMI_Status".Status.ZoneStatusIndex].StartPos;
END_REGION

REGION Network 46
   RUNG wire#powerrail
      Move(in := "EMS".Zone["DB401_HMI_Status".Status.ZoneStatusIndex].EndPos, out1 => "DB401_HMI_Status".ZoneStatus.ZoneEndPosition)
   END_RUNG
   // the same network as SCL:
   "DB401_HMI_Status".ZoneStatus.ZoneEndPosition := "EMS".Zone["DB401_HMI_Status".Status.ZoneStatusIndex].EndPos;
END_REGION

REGION Network 47
   RUNG wire#powerrail
      Move(in := "EMS".Zone["DB401_HMI_Status".Status.ZoneStatusIndex].PrevZone, out1 => "DB401_HMI_Status".ZoneStatus.PrevZoneNumber)
   END_RUNG
   // the same network as SCL:
   "DB401_HMI_Status".ZoneStatus.PrevZoneNumber := "EMS".Zone["DB401_HMI_Status".Status.ZoneStatusIndex].PrevZone;
END_REGION

REGION Network 48
   RUNG wire#powerrail
      Move(in := "EMS".Zone["DB401_HMI_Status".Status.ZoneStatusIndex].NextZone, out1 => "DB401_HMI_Status".ZoneStatus.NextZoneNumber)
   END_RUNG
   // the same network as SCL:
   "DB401_HMI_Status".ZoneStatus.NextZoneNumber := "EMS".Zone["DB401_HMI_Status".Status.ZoneStatusIndex].NextZone;
END_REGION

REGION Network 49
   RUNG wire#powerrail
      Move(in := "EMS".Zone["DB401_HMI_Status".Status.ZoneStatusIndex].SpeedZoneStart, out1 => "DB401_HMI_Status".ZoneStatus.SpeedZoneStartPos)
   END_RUNG
   // the same network as SCL:
   "DB401_HMI_Status".ZoneStatus.SpeedZoneStartPos := "EMS".Zone["DB401_HMI_Status".Status.ZoneStatusIndex].SpeedZoneStart;
END_REGION

REGION Network 50
   RUNG wire#powerrail
      Move(in := "EMS".Zone["DB401_HMI_Status".Status.ZoneStatusIndex].SpeedZoneEnd, out1 => "DB401_HMI_Status".ZoneStatus.SpeedZoneEndPos)
   END_RUNG
   // the same network as SCL:
   "DB401_HMI_Status".ZoneStatus.SpeedZoneEndPos := "EMS".Zone["DB401_HMI_Status".Status.ZoneStatusIndex].SpeedZoneEnd;
END_REGION

REGION Network 51
